REGION Network 12: Lowest Value of 2
   RUNG wire#powerrail
      Contact( #HMI.Alarms.oneTxFaulted )
      I_Contact( #HMI.Alarms.twoTxFaulted )
      { S7_Templates := "SrcType := Int" } EQ_Contact(in1 := #HMI.Control.failMode, in2 := 7)
      Move(in := #lowest, out1 => #activeValue)
   END_RUNG
   // the same network as SCL:
   IF #HMI.Alarms.oneTxFaulted AND NOT #HMI.Alarms.twoTxFaulted AND (#HMI.Control.failMode = 7) THEN
       #activeValue := #lowest;
   END_IF;
END_REGION

REGION Network 13: Average Value
   RUNG wire#powerrail
      Contact( #fault3 )
      { S7_Templates := "SrcType := Real"; S7_Expression := "(IN1+IN2)/IN3" } Calculate(in1 := #analog1, in2 := #analog2, in3 := 2.0, out => #average)
   END_RUNG
   RUNG wire#powerrail
      Contact( #fault2 )
      { S7_Templates := "SrcType := Real"; S7_Expression := "(IN1+IN2)/IN3" } Calculate(in1 := #analog1, in2 := #analog3, in3 := 2.0, out => #average)
   END_RUNG
   RUNG wire#powerrail
      Contact( #fault1 )
      { S7_Templates := "SrcType := Real"; S7_Expression := "(IN1+IN2)/IN3" } Calculate(in1 := #analog3, in2 := #analog2, in3 := 2.0, out => #average)
   END_RUNG
   RUNG wire#powerrail
      I_Contact( #fault1 )
      I_Contact( #fault2 )
      I_Contact( #fault3 )
      { S7_Templates := "SrcType := Real"; S7_Expression := "(IN1+IN2+IN3)/IN4" } Calculate(in1 := #analog1, in2 := #analog2, in3 := #analog3, in4 := 3.0, out => #average)
   END_RUNG
   // the same network as SCL:
   IF #fault3 THEN #average := (#analog1+#analog2)/2.0; END_IF;
   IF #fault2 THEN #average := (#analog1+#analog3)/2.0; END_IF;
   IF #fault1 THEN #average := (#analog3+#analog2)/2.0; END_IF;
   IF NOT #fault1 AND NOT #fault2 AND NOT #fault3 THEN #average := (#analog1+#analog2+#analog3)/3.0; END_IF;
END_REGION

REGION Network 14: Average of 3 values
   RUNG wire#powerrail
      { S7_Templates := "SrcType := Int" } EQ_Contact(in1 := #HMI.Control.mode, in2 := 4)
      wire#w1
      Move(in := #average, out1 => #activeValue)
   END_RUNG
   RUNG wire#powerrail
      Contact( #HMI.Alarms.oneTxFaulted )
      I_Contact( #HMI.Alarms.twoTxFaulted )
      { S7_Templates := "SrcType := Int" } EQ_Contact(in1 := #HMI.Control.failMode, in2 := 4)
   END_RUNG wire#w1
   // the same network as SCL:
   IF (#HMI.Control.mode = 4) OR (#HMI.Alarms.oneTxFaulted AND NOT #HMI.Alarms.twoTxFaulted AND (#HMI.Control.failMode = 4)) THEN
       #activeValue := #average;
   END_IF;
END_REGION

REGION Network 15: HH Voting Value 1
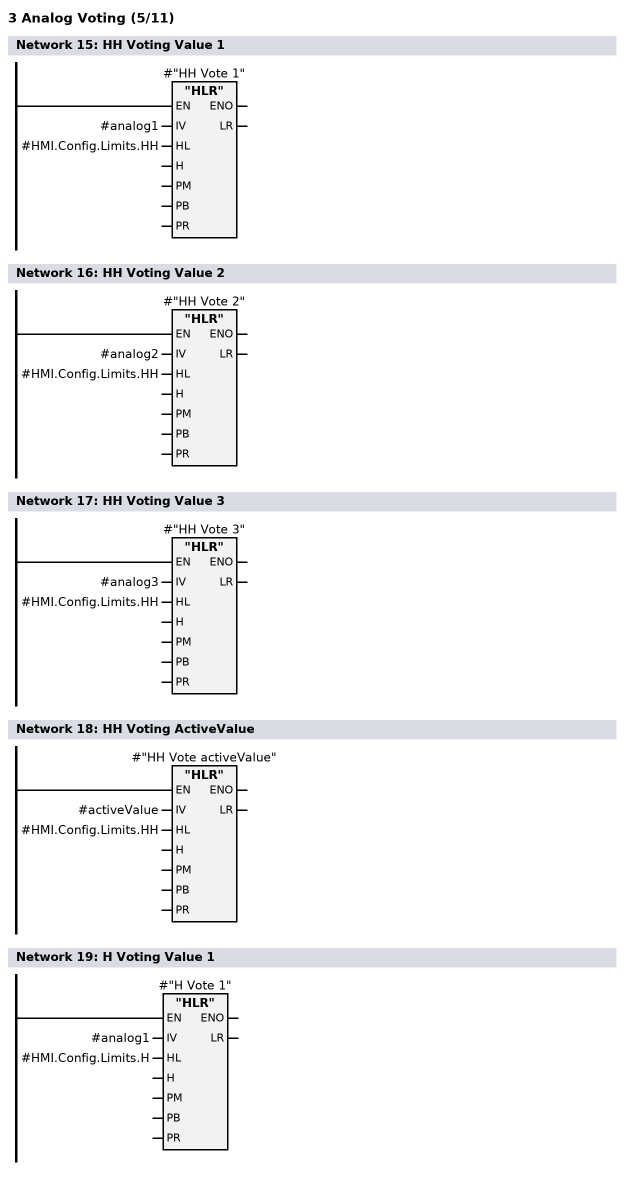
   RUNG wire#powerrail
      #"HH Vote 1"(IV := #analog1, HL := #HMI.Config.Limits.HH, H :=, PM :=, PB :=, PR :=, LR =>)
   END_RUNG
   // the same network as SCL:
   #"HH Vote 1"(IV := #analog1, HL := #HMI.Config.Limits.HH);   // "HLR"
END_REGION

REGION Network 16: HH Voting Value 2
   RUNG wire#powerrail
      #"HH Vote 2"(IV := #analog2, HL := #HMI.Config.Limits.HH, H :=, PM :=, PB :=, PR :=, LR =>)
   END_RUNG
   // the same network as SCL:
   #"HH Vote 2"(IV := #analog2, HL := #HMI.Config.Limits.HH);   // "HLR"
END_REGION

REGION Network 17: HH Voting Value 3
   RUNG wire#powerrail
      #"HH Vote 3"(IV := #analog3, HL := #HMI.Config.Limits.HH, H :=, PM :=, PB :=, PR :=, LR =>)
   END_RUNG
   // the same network as SCL:
   #"HH Vote 3"(IV := #analog3, HL := #HMI.Config.Limits.HH);   // "HLR"
END_REGION

REGION Network 18: HH Voting ActiveValue
   RUNG wire#powerrail
      #"HH Vote activeValue"(IV := #activeValue, HL := #HMI.Config.Limits.HH, H :=, PM :=, PB :=, PR :=, LR =>)
   END_RUNG
   // the same network as SCL:
   #"HH Vote activeValue"(IV := #activeValue, HL := #HMI.Config.Limits.HH);   // "HLR"
END_REGION

REGION Network 19: H Voting Value 1
   RUNG wire#powerrail
      #"H Vote 1"(IV := #analog1, HL := #HMI.Config.Limits.H, H :=, PM :=, PB :=, PR :=, LR =>)
   END_RUNG
   // the same network as SCL:
   #"H Vote 1"(IV := #analog1, HL := #HMI.Config.Limits.H);   // "HLR"
END_REGION

REGION Network 20: H Voting Value 2
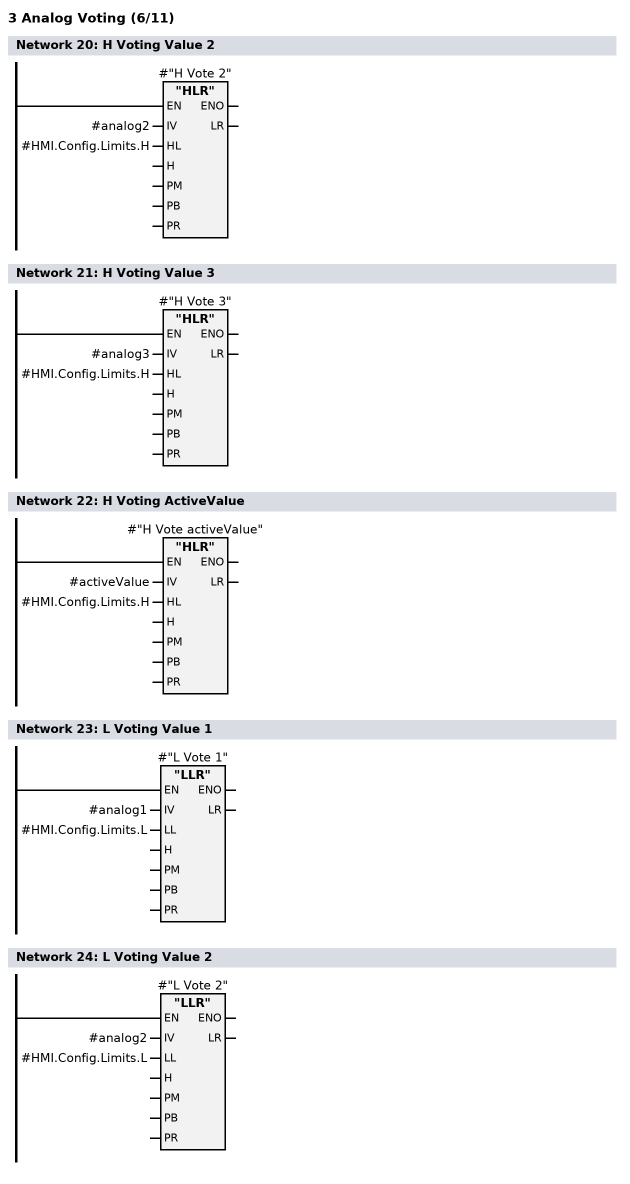
   RUNG wire#powerrail
      #"H Vote 2"(IV := #analog2, HL := #HMI.Config.Limits.H, H :=, PM :=, PB :=, PR :=, LR =>)
   END_RUNG
   // the same network as SCL:
   #"H Vote 2"(IV := #analog2, HL := #HMI.Config.Limits.H);   // "HLR"
END_REGION

REGION Network 21: H Voting Value 3
   RUNG wire#powerrail
      #"H Vote 3"(IV := #analog3, HL := #HMI.Config.Limits.H, H :=, PM :=, PB :=, PR :=, LR =>)
   END_RUNG
   // the same network as SCL:
   #"H Vote 3"(IV := #analog3, HL := #HMI.Config.Limits.H);   // "HLR"
END_REGION

REGION Network 22: H Voting ActiveValue
   RUNG wire#powerrail
      #"H Vote activeValue"(IV := #activeValue, HL := #HMI.Config.Limits.H, H :=, PM :=, PB :=, PR :=, LR =>)
   END_RUNG
   // the same network as SCL:
   #"H Vote activeValue"(IV := #activeValue, HL := #HMI.Config.Limits.H);   // "HLR"
END_REGION

REGION Network 23: L Voting Value 1
   RUNG wire#powerrail
      #"L Vote 1"(IV := #analog1, LL := #HMI.Config.Limits.L, H :=, PM :=, PB :=, PR :=, LR =>)
   END_RUNG
   // the same network as SCL:
   #"L Vote 1"(IV := #analog1, LL := #HMI.Config.Limits.L);   // "LLR"
END_REGION

REGION Network 24: L Voting Value 2
   RUNG wire#powerrail
      #"L Vote 2"(IV := #analog2, LL := #HMI.Config.Limits.L, H :=, PM :=, PB :=, PR :=, LR =>)
   END_RUNG
   // the same network as SCL:
   #"L Vote 2"(IV := #analog2, LL := #HMI.Config.Limits.L);   // "LLR"
END_REGION

REGION Network 25: L Voting Value 3
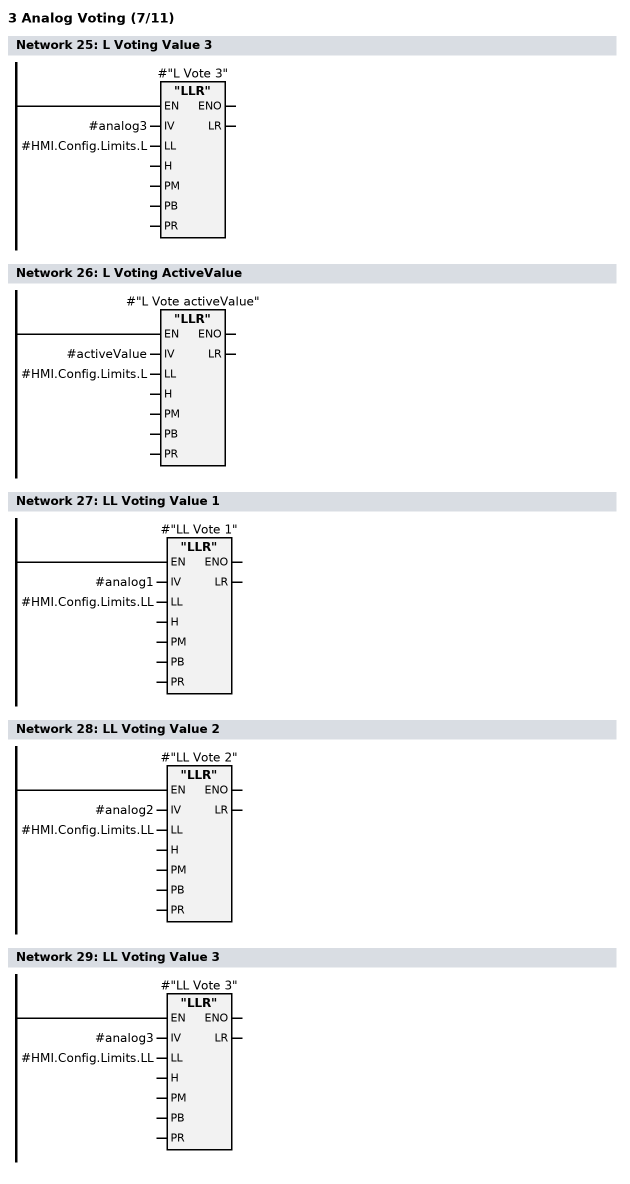
   RUNG wire#powerrail
      #"L Vote 3"(IV := #analog3, LL := #HMI.Config.Limits.L, H :=, PM :=, PB :=, PR :=, LR =>)
   END_RUNG
   // the same network as SCL:
   #"L Vote 3"(IV := #analog3, LL := #HMI.Config.Limits.L);   // "LLR"
END_REGION

REGION Network 26: L Voting ActiveValue
   RUNG wire#powerrail
      #"L Vote activeValue"(IV := #activeValue, LL := #HMI.Config.Limits.L, H :=, PM :=, PB :=, PR :=, LR =>)
   END_RUNG
   // the same network as SCL:
   #"L Vote activeValue"(IV := #activeValue, LL := #HMI.Config.Limits.L);   // "LLR"
END_REGION

REGION Network 27: LL Voting Value 1
   RUNG wire#powerrail
      #"LL Vote 1"(IV := #analog1, LL := #HMI.Config.Limits.LL, H :=, PM :=, PB :=, PR :=, LR =>)
   END_RUNG
   // the same network as SCL:
   #"LL Vote 1"(IV := #analog1, LL := #HMI.Config.Limits.LL);   // "LLR"
END_REGION

REGION Network 28: LL Voting Value 2
   RUNG wire#powerrail
      #"LL Vote 2"(IV := #analog2, LL := #HMI.Config.Limits.LL, H :=, PM :=, PB :=, PR :=, LR =>)
   END_RUNG
   // the same network as SCL:
   #"LL Vote 2"(IV := #analog2, LL := #HMI.Config.Limits.LL);   // "LLR"
END_REGION

REGION Network 29: LL Voting Value 3
   RUNG wire#powerrail
      #"LL Vote 3"(IV := #analog3, LL := #HMI.Config.Limits.LL, H :=, PM :=, PB :=, PR :=, LR =>)
   END_RUNG
   // the same network as SCL:
   #"LL Vote 3"(IV := #analog3, LL := #HMI.Config.Limits.LL);   // "LLR"
END_REGION

REGION Network 30: LL Voting ActiveValue
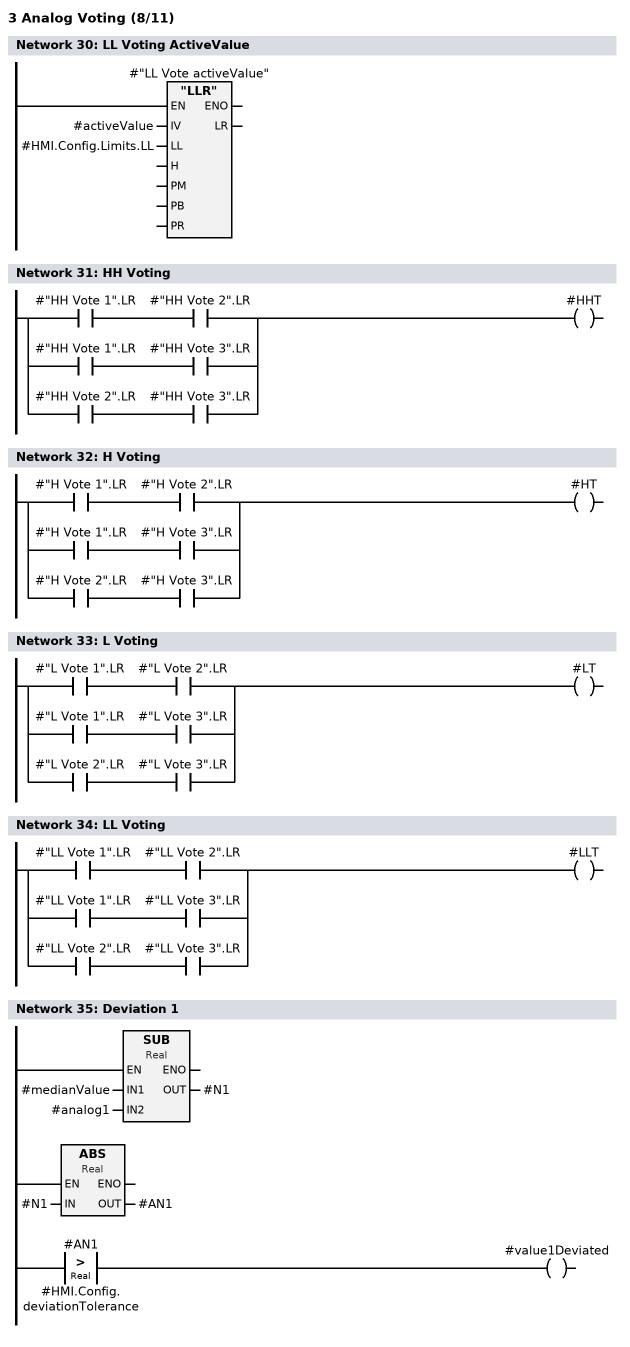
   RUNG wire#powerrail
      #"LL Vote activeValue"(IV := #activeValue, LL := #HMI.Config.Limits.LL, H :=, PM :=, PB :=, PR :=, LR =>)
   END_RUNG
   // the same network as SCL:
   #"LL Vote activeValue"(IV := #activeValue, LL := #HMI.Config.Limits.LL);   // "LLR"
END_REGION

REGION Network 31: HH Voting
   RUNG wire#powerrail
      Contact( #"HH Vote 1".LR )
      Contact( #"HH Vote 2".LR )
      wire#w1
      Coil( #HHT )
   END_RUNG
   RUNG wire#powerrail
      Contact( #"HH Vote 1".LR )
      Contact( #"HH Vote 3".LR )
   END_RUNG wire#w1
   RUNG wire#powerrail
      Contact( #"HH Vote 2".LR )
      Contact( #"HH Vote 3".LR )
   END_RUNG wire#w1
   // the same network as SCL:
   #HHT := (#"HH Vote 1".LR AND #"HH Vote 2".LR) OR (#"HH Vote 1".LR AND #"HH Vote 3".LR) OR (#"HH Vote 2".LR AND #"HH Vote 3".LR);
END_REGION

REGION Network 32: H Voting
   RUNG wire#powerrail
      Contact( #"H Vote 1".LR )
      Contact( #"H Vote 2".LR )
      wire#w1
      Coil( #HT )
   END_RUNG
   RUNG wire#powerrail
      Contact( #"H Vote 1".LR )
      Contact( #"H Vote 3".LR )
   END_RUNG wire#w1
   RUNG wire#powerrail
      Contact( #"H Vote 2".LR )
      Contact( #"H Vote 3".LR )
   END_RUNG wire#w1
   // the same network as SCL:
   #HT := (#"H Vote 1".LR AND #"H Vote 2".LR) OR (#"H Vote 1".LR AND #"H Vote 3".LR) OR (#"H Vote 2".LR AND #"H Vote 3".LR);
END_REGION

REGION Network 33: L Voting
   RUNG wire#powerrail
      Contact( #"L Vote 1".LR )
      Contact( #"L Vote 2".LR )
      wire#w1
      Coil( #LT )
   END_RUNG
   RUNG wire#powerrail
      Contact( #"L Vote 1".LR )
      Contact( #"L Vote 3".LR )
   END_RUNG wire#w1
   RUNG wire#powerrail
      Contact( #"L Vote 2".LR )
      Contact( #"L Vote 3".LR )
   END_RUNG wire#w1
   // the same network as SCL:
   #LT := (#"L Vote 1".LR AND #"L Vote 2".LR) OR (#"L Vote 1".LR AND #"L Vote 3".LR) OR (#"L Vote 2".LR AND #"L Vote 3".LR);
END_REGION

REGION Network 34: LL Voting
   RUNG wire#powerrail
      Contact( #"LL Vote 1".LR )
      Contact( #"LL Vote 2".LR )
      wire#w1
      Coil( #LLT )
   END_RUNG
   RUNG wire#powerrail
      Contact( #"LL Vote 1".LR )
      Contact( #"LL Vote 3".LR )
   END_RUNG wire#w1
   RUNG wire#powerrail
      Contact( #"LL Vote 2".LR )
      Contact( #"LL Vote 3".LR )
   END_RUNG wire#w1
   // the same network as SCL:
   #LLT := (#"LL Vote 1".LR AND #"LL Vote 2".LR) OR (#"LL Vote 1".LR AND #"LL Vote 3".LR) OR (#"LL Vote 2".LR AND #"LL Vote 3".LR);
END_REGION

REGION Network 35: Deviation 1
   RUNG wire#powerrail
      { S7_Templates := "SrcType := Real"; S7_GenerateENO := "TRUE" } Sub(in1 := #medianValue, in2 := #analog1, out => #N1)
   END_RUNG
   RUNG wire#powerrail
      { S7_Templates := "SrcType := Real"; S7_GenerateENO := "TRUE" } Abs(in := #N1, out => #AN1)
   END_RUNG
   RUNG wire#powerrail
      { S7_Templates := "SrcType := Real" } GT_Contact(in1 := #AN1, in2 := #HMI.Config.deviationTolerance)
      Coil( #value1Deviated )
   END_RUNG
   // the same network as SCL:
   #N1 := #medianValue - #analog1;
   #AN1 := ABS(#N1);
   #value1Deviated := #AN1 > #HMI.Config.deviationTolerance;
END_REGION

REGION Network 36: Deviation 2
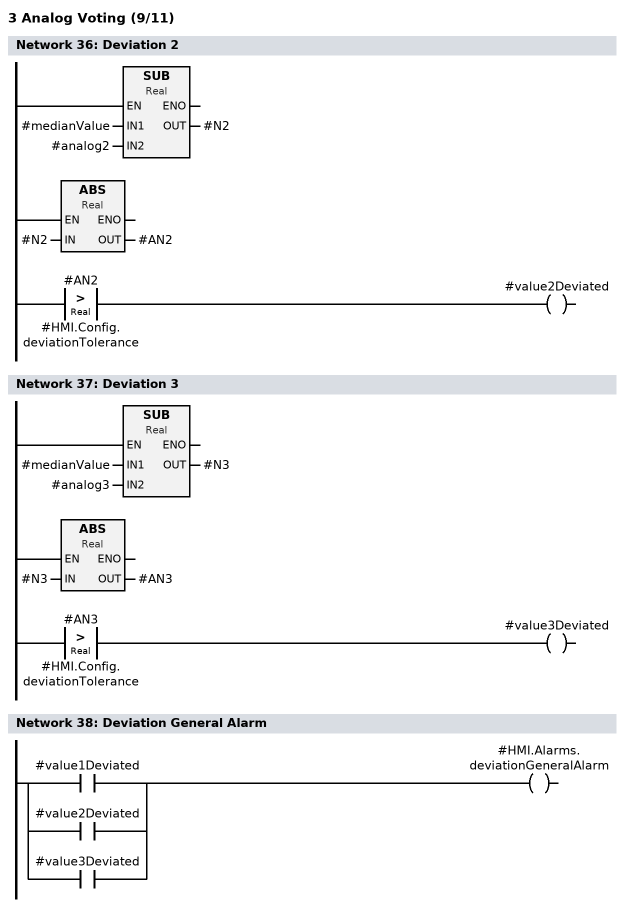
   RUNG wire#powerrail
      { S7_Templates := "SrcType := Real"; S7_GenerateENO := "TRUE" } Sub(in1 := #medianValue, in2 := #analog2, out => #N2)
   END_RUNG
   RUNG wire#powerrail
      { S7_Templates := "SrcType := Real"; S7_GenerateENO := "TRUE" } Abs(in := #N2, out => #AN2)
   END_RUNG
   RUNG wire#powerrail
      { S7_Templates := "SrcType := Real" } GT_Contact(in1 := #AN2, in2 := #HMI.Config.deviationTolerance)
      Coil( #value2Deviated )
   END_RUNG
   // the same network as SCL:
   #N2 := #medianValue - #analog2;
   #AN2 := ABS(#N2);
   #value2Deviated := #AN2 > #HMI.Config.deviationTolerance;
END_REGION

REGION Network 37: Deviation 3
   RUNG wire#powerrail
      { S7_Templates := "SrcType := Real"; S7_GenerateENO := "TRUE" } Sub(in1 := #medianValue, in2 := #analog3, out => #N3)
   END_RUNG
   RUNG wire#powerrail
      { S7_Templates := "SrcType := Real"; S7_GenerateENO := "TRUE" } Abs(in := #N3, out => #AN3)
   END_RUNG
   RUNG wire#powerrail
      { S7_Templates := "SrcType := Real" } GT_Contact(in1 := #AN3, in2 := #HMI.Config.deviationTolerance)
      Coil( #value3Deviated )
   END_RUNG
   // the same network as SCL:
   #N3 := #medianValue - #analog3;
   #AN3 := ABS(#N3);
   #value3Deviated := #AN3 > #HMI.Config.deviationTolerance;
END_REGION

REGION Network 38: Deviation General Alarm
   RUNG wire#powerrail
      Contact( #value1Deviated )
      wire#w1
      Coil( #HMI.Alarms.deviationGeneralAlarm )
   END_RUNG
   RUNG wire#powerrail
      Contact( #value2Deviated )
   END_RUNG wire#w1
   RUNG wire#powerrail
      Contact( #value3Deviated )
   END_RUNG wire#w1
   // the same network as SCL:
   #HMI.Alarms.deviationGeneralAlarm := #value1Deviated OR #value2Deviated OR #value3Deviated;
END_REGION

REGION Network 39: Master Trip
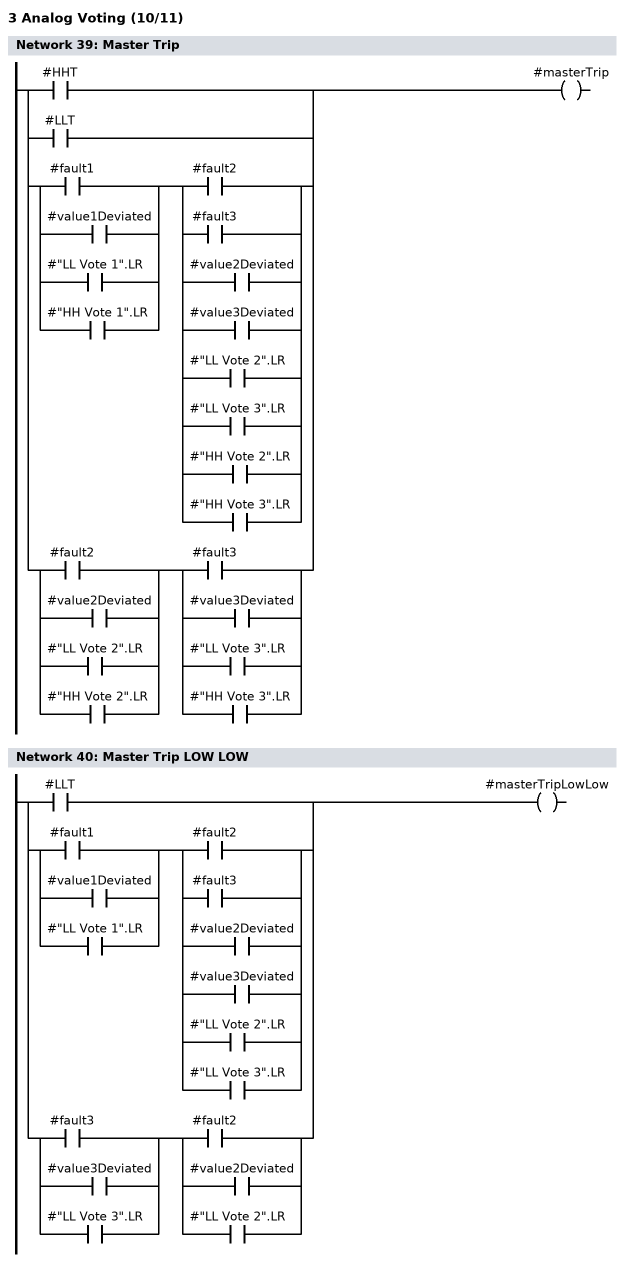
   RUNG wire#powerrail
      Contact( #HHT )
      wire#w1
      Coil( #masterTrip )
   END_RUNG
   RUNG wire#powerrail
      Contact( #LLT )
   END_RUNG wire#w1
   RUNG wire#powerrail
      Contact( #fault1 )
      wire#w2
      Contact( #fault2 )
   END_RUNG wire#w1
   RUNG wire#powerrail
      Contact( #value1Deviated )
   END_RUNG wire#w2
   RUNG wire#powerrail
      Contact( #"LL Vote 1".LR )
   END_RUNG wire#w2
   RUNG wire#powerrail
      Contact( #"HH Vote 1".LR )
   END_RUNG wire#w2
   RUNG wire#w2
      Contact( #fault3 )
   END_RUNG wire#w1
   RUNG wire#w2
      Contact( #value2Deviated )
   END_RUNG wire#w1
   RUNG wire#w2
      Contact( #value3Deviated )
   END_RUNG wire#w1
   RUNG wire#w2
      Contact( #"LL Vote 2".LR )
   END_RUNG wire#w1
   RUNG wire#w2
      Contact( #"LL Vote 3".LR )
   END_RUNG wire#w1
   RUNG wire#w2
      Contact( #"HH Vote 2".LR )
   END_RUNG wire#w1
   RUNG wire#w2
      Contact( #"HH Vote 3".LR )
   END_RUNG wire#w1
   RUNG wire#powerrail
      Contact( #fault2 )
      wire#w3
      Contact( #fault3 )
   END_RUNG wire#w1
   RUNG wire#powerrail
      Contact( #value2Deviated )
   END_RUNG wire#w3
   RUNG wire#powerrail
      Contact( #"LL Vote 2".LR )
   END_RUNG wire#w3
   RUNG wire#powerrail
      Contact( #"HH Vote 2".LR )
   END_RUNG wire#w3
   RUNG wire#w3
      Contact( #value3Deviated )
   END_RUNG wire#w1
   RUNG wire#w3
      Contact( #"LL Vote 3".LR )
   END_RUNG wire#w1
   RUNG wire#w3
      Contact( #"HH Vote 3".LR )
   END_RUNG wire#w1
   // the same network as SCL:
   #masterTrip := #HHT OR #LLT OR ((#fault1 OR #value1Deviated OR #"LL Vote 1".LR OR #"HH Vote 1".LR) AND (#fault2 OR #fault3 OR #value2Deviated OR #value3Deviated OR #"LL Vote 2".LR OR #"LL Vote 3".LR OR #"HH Vote 2".LR OR #"HH Vote 3".LR)) OR ((#fault2 OR #value2Deviated OR #"LL Vote 2".LR OR #"HH Vote 2".LR) AND (#fault3 OR #value3Deviated OR #"LL Vote 3".LR OR #"HH Vote 3".LR));
END_REGION

REGION Network 40: Master Trip LOW LOW
   RUNG wire#powerrail
      Contact( #LLT )
      wire#w1
      Coil( #masterTripLowLow )
   END_RUNG
   RUNG wire#powerrail
      Contact( #fault1 )
      wire#w2
      Contact( #fault2 )
   END_RUNG wire#w1
   RUNG wire#powerrail
      Contact( #value1Deviated )
   END_RUNG wire#w2
   RUNG wire#powerrail
      Contact( #"LL Vote 1".LR )
   END_RUNG wire#w2
   RUNG wire#w2
      Contact( #fault3 )
   END_RUNG wire#w1
   RUNG wire#w2
      Contact( #value2Deviated )
   END_RUNG wire#w1
   RUNG wire#w2
      Contact( #value3Deviated )
   END_RUNG wire#w1
   RUNG wire#w2
      Contact( #"LL Vote 2".LR )
   END_RUNG wire#w1
   RUNG wire#w2
      Contact( #"LL Vote 3".LR )
   END_RUNG wire#w1
   RUNG wire#powerrail
      Contact( #fault3 )
      wire#w3
      Contact( #fault2 )
   END_RUNG wire#w1
   RUNG wire#powerrail
      Contact( #value3Deviated )
   END_RUNG wire#w3
   RUNG wire#powerrail
      Contact( #"LL Vote 3".LR )
   END_RUNG wire#w3
   RUNG wire#w3
      Contact( #value2Deviated )
   END_RUNG wire#w1
   RUNG wire#w3
      Contact( #"LL Vote 2".LR )
   END_RUNG wire#w1
   // the same network as SCL:
   #masterTripLowLow := #LLT OR ((#fault1 OR #value1Deviated OR #"LL Vote 1".LR) AND (#fault2 OR #fault3 OR #value2Deviated OR #value3Deviated OR #"LL Vote 2".LR OR #"LL Vote 3".LR)) OR ((#fault3 OR #value3Deviated OR #"LL Vote 3".LR) AND (#fault2 OR #value2Deviated OR #"LL Vote 2".LR));
END_REGION

REGION Network 41: Master Trip HIGH HIGH
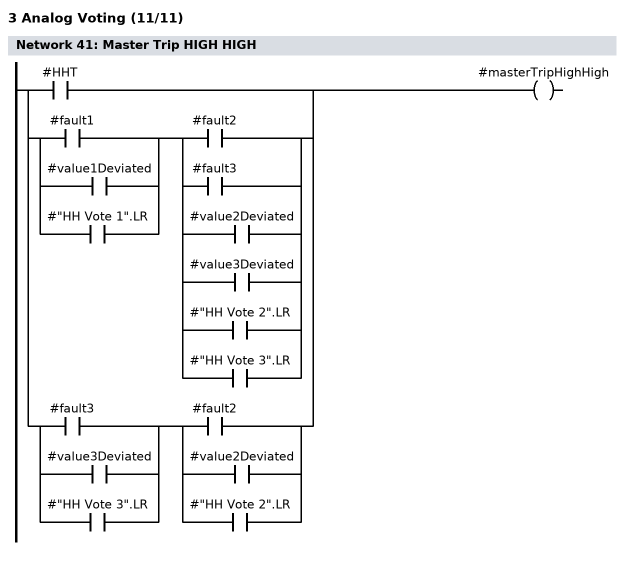
   RUNG wire#powerrail
      Contact( #HHT )
      wire#w1
      Coil( #masterTripHighHigh )
   END_RUNG
   RUNG wire#powerrail
      Contact( #fault1 )
      wire#w2
      Contact( #fault2 )
   END_RUNG wire#w1
   RUNG wire#powerrail
      Contact( #value1Deviated )
   END_RUNG wire#w2
   RUNG wire#powerrail
      Contact( #"HH Vote 1".LR )
   END_RUNG wire#w2
   RUNG wire#w2
      Contact( #fault3 )
   END_RUNG wire#w1
   RUNG wire#w2
      Contact( #value2Deviated )
   END_RUNG wire#w1
   RUNG wire#w2
      Contact( #value3Deviated )
   END_RUNG wire#w1
   RUNG wire#w2
      Contact( #"HH Vote 2".LR )
   END_RUNG wire#w1
   RUNG wire#w2
      Contact( #"HH Vote 3".LR )
   END_RUNG wire#w1
   RUNG wire#powerrail
      Contact( #fault3 )
      wire#w3
      Contact( #fault2 )
   END_RUNG wire#w1
   RUNG wire#powerrail
      Contact( #value3Deviated )
   END_RUNG wire#w3
   RUNG wire#powerrail
      Contact( #"HH Vote 3".LR )
   END_RUNG wire#w3
   RUNG wire#w3
      Contact( #value2Deviated )
   END_RUNG wire#w1
   RUNG wire#w3
      Contact( #"HH Vote 2".LR )
   END_RUNG wire#w1
   // the same network as SCL:
   #masterTripHighHigh := #HHT OR ((#fault1 OR #value1Deviated OR #"HH Vote 1".LR) AND (#fault2 OR #fault3 OR #value2Deviated OR #value3Deviated OR #"HH Vote 2".LR OR #"HH Vote 3".LR)) OR ((#fault3 OR #value3Deviated OR #"HH Vote 3".LR) AND (#fault2 OR #value2Deviated OR #"HH Vote 2".LR));
END_REGION
END_FUNCTION_BLOCK

FUNCTION_BLOCK "TX-AI"   // FB804, LAD
TITLE = SSAC Analog Trasmitter Function Block
{ S7_Optimized_Access := 'TRUE' }
VERSION : 1.0
// Default mode 0 starts at  network 6
   VAR_INPUT
      Mode : Int;   // TX Mode - 0 = 4-20 mA / 1 = Int Math (RTD/TC) / 2 = Real Input Conversion / 3 = SQRT / 5 = Simulated Transmitter Value / 6 = Vortex Flow Transmitters
      RAIVI : Int;   // Raw Analog Input Value INT
      RAIVR : Real;   // Raw Analog Input Value REAL
      EnableHighAlarms : Bool := True;
      EnableLowAlarms : Bool := True;
      "TI Fail" : Bool;
   END_VAR
   VAR_OUTPUT
      SAI : Real;   // Compensated Scaled Analog Value
   END_VAR
   VAR
      HMI : Struct   // Alarms
         Status : Struct
            USAV : Real;   // Uncompensated Scaled Analog Value
            TCV : Real;   // Temperature Compensation Value
            PCV : Real;   // Pressure Compensation Value
            NV : Real;   // Normalized Value
         END_STRUCT;
         Alarm : Struct
            Alarms : Word;
         END_STRUCT;
         Diag : Struct   // Diagnostics
            SV : Real;   // Simulation Value
         END_STRUCT;
      END_STRUCT;
   END_VAR
   VAR RETAIN
      Retain : Struct
         HMI : Struct
            Config : Struct   // Settings
               RIMXV : Real := 27648.0;   // Raw Input Maximum Value (Used for Sqrt)
               RIMNV : Real;   // Raw Input Minimum Value (Used for Sqrt)
               ESMXV : Real := 100.0;   // Engineering/Scaled Maximum Value
               ESMNV : Real;   // Engineering/Scaled Minimum Value
               COV : Bool;   // Clamp Output Value
               OV : Real;   // Offset Value
               SAM : Bool;   // Substitution Activation Mode
               SAV : Real := -999999.0;   // Substitution Value during a limit input value trip
               CE : Struct   // Compensation Equation
                  TC : Real := 460.0;   // Temperature Constant
                  PC : Real := 14.7;   // Pressure Constant
                  TR : Real := 1.0;   // Temperature Reference
                  TA : Real := 1.0;   // Temperature Actual
                  PR : Real := 1.0;   // Pressure Reference
                  PA : Real := 1.0;   // Pressure Actual
               END_STRUCT;
               SP : Struct   // Setpoints
                  Limits : Struct
                     HHH : Real := 95.0;   // HHH Limit Setpoint
                     HH : Real := 90.0;   // HH Limit Setpoint
                     H : Real := 80.0;   // HH Limit Setpoint
                     L : Real := 20.0;   // L Limit Setpoint
                     LL : Real := 10.0;   // LL Limit Setpoint
                     LLL : Real := 5.0;   // LLL Limit Setpoint
                     "OR" : Real := 5.0;   // Over range value
                     UR : Real := 5.0;   // Under range value
                  END_STRUCT;
                  HYS : Struct   // Hysteresis
                     Global : Real;   // Hysteresis global value, only valid when greater than or equal to 0
                     HHH : Real := 1.0;   // Hysteresis Setpoint - High High High
                     HH : Real := 1.0;   // Hysteresis Setpoint - High High
                     H : Real := 1.0;   // Hysteresis Setpoint - High
                     L : Real := 1.0;   // Hysteresis Setpoint - Low
                     LL : Real := 1.0;   // Hysteresis Setpoint - Low Low
                     LLL : Real := 1.0;   // Hysteresis Setpoint - Low Low Low
                     "OR" : Real := 1.0;   // Hysteresis Setpoint - Over Range
                     UR : Real := 1.0;   // Hysteresis Setpoint - Under Range
                  END_STRUCT;
                  SUB_ON : Bool;   // Substitution Activation
               END_STRUCT;
               PT : Struct   // Setpoints
                  HLD : Struct   // Hold
                     Global : Time;   // Hold PT global value, only valid when not equal to 0
                     AHHH : Time := t#5s;   // Alarm Debounce
                     AHH : Time := t#5s;   // Alarm Debounce
                     AH : Time := t#5s;   // Alarm Debounce
                     AL : Time := t#5s;   // Alarm Debounce
                     ALL : Time := t#5s;   // Alarm Debounce
                     ALLL : Time := t#5s;   // Alarm Debounce
                     "OR" : Time := t#5s;   // Over range hold
                     UR : Time := t#5s;   // Under range hold
                  END_STRUCT;
                  DBNC : Struct   // Debounce
                     Global : Time;   // Debounce PT global value, only valid when not equal to 0
                     AHHH : Time := t#5s;   // Alarm Debounce
                     AHH : Time := t#5s;   // Alarm Debounce
                     AH : Time := t#5s;   // Alarm Debounce
                     AL : Time := t#5s;   // Alarm Debounce
                     ALL : Time := t#5s;   // Alarm Debounce
                     ALLL : Time := t#5s;   // Alarm Debounce
                     "OR" : Time := t#5s;   // Over range debounce
                     UR : Time := t#5s;   // Under range debounce
                  END_STRUCT;
               END_STRUCT;
               Alarms : Word := 16#01FF;
            END_STRUCT;
         END_STRUCT;
      END_STRUCT;
   END_VAR
   VAR
      Admin : Struct   // Admin configurations
         SCL : Struct   // Scale Values
            RDP : Real := 10.0;   // RTD Decimal Places
            RRIMD : Real := 1.0;   // Raw Real input Math divider
            "OR" : Real;   // Over Range Value
            UR : Real;   // Under Range Value
            SAIV : Real;   // Scaled Analog Input Value
         END_STRUCT;
         HYS : Struct   // Hysteresis - Computed Values
            "OR" : Real;   // Hysteresis Value - Over Range
            UR : Real;   // Hysteresis Value - Under Range
         END_STRUCT;
      END_STRUCT;
      Alarms : Struct
         HighHighHigh : Bool;
         HighHigh : Bool;
         High : Bool;
         Low : Bool;
         LowLow : Bool;
         LowLowLow : Bool;
         TransmitterFault : Bool;
         UnderRange : Bool;
         OverRange : Bool;
      END_STRUCT;
      Timers : Struct
         OR_DB : TON_TIME;   // Over Range Debounce
         UR_DB : TON_TIME;   // Under Range DB
         OR_HLD : TOF_TIME;   // Over Range Hold
         UR_HLD : TOF_TIME;   // Under Range Hold
         DBNC : Struct
            HHH : TON_TIME;
            HH : TON_TIME;
            H : TON_TIME;
            L : TON_TIME;
            LL : TON_TIME;
            LLL : TON_TIME;
         END_STRUCT;
         HOLD : Struct
            HHH : TOF_TIME;
            HH : TOF_TIME;
            H : TOF_TIME;
            L : TOF_TIME;
            LL : TOF_TIME;
            LLL : TOF_TIME;
         END_STRUCT;
      END_STRUCT;
      molActual : Real := 1.0;
      molDesign : Real := 1.0;
   END_VAR
   VAR_TEMP
      SRV : Real;
      RAIDI : DInt;   // Raw Analog Input DINT
      RAIR : Real;   // Raw Analog Input REAL
      RAIAV : Real;   // Raw Analog Input Absolute Value
      RAIVS : Real;   // Raw Analog Input Value Scaler
      TCRE : Real;   // Temperature Compensation Reference Equation
      TCAE : Real;   // Temperature Compensation Actual Equation
      PCRE : Real;   // Pressure Compensation Reference Equation
      PCAE : Real;   // Pressure Compensation Actual Equation
      TPCV : Real;   // Temperature Pressure Compensation Value
      MWCV : Real;   // Mol Weight Compensation Value
      TPMCV : Real;   // Temperature Pressure Mol Compensation Value
      sqrtSaiv : Real;   // SCALED ANALOG INT VALUE TO BE SQRT'D
      rawValue : Int;
      dummy : Bool;
      sqrt01 : Real;
      RAIVR_1 : DInt;
      RAIVR_1_1 : Real;
      ValuePerPoint : Real;
      ValueAddRaw : Real;
      "DBNC.SP" : Struct
         HHH : Real;
         HH : Real;
         H : Real;
         L : Real;
         LL : Real;
         LLL : Real;
      END_STRUCT;
   END_VAR
   VAR_TEMP   // added for the SCL form of the ladder/FBD networks
      _w1 : Bool;
      _w2 : Bool;
   END_VAR
BEGIN

REGION Network 1: Transmitter Mode 1 = Int Math or RTD
   // MD1 Jump to network 9
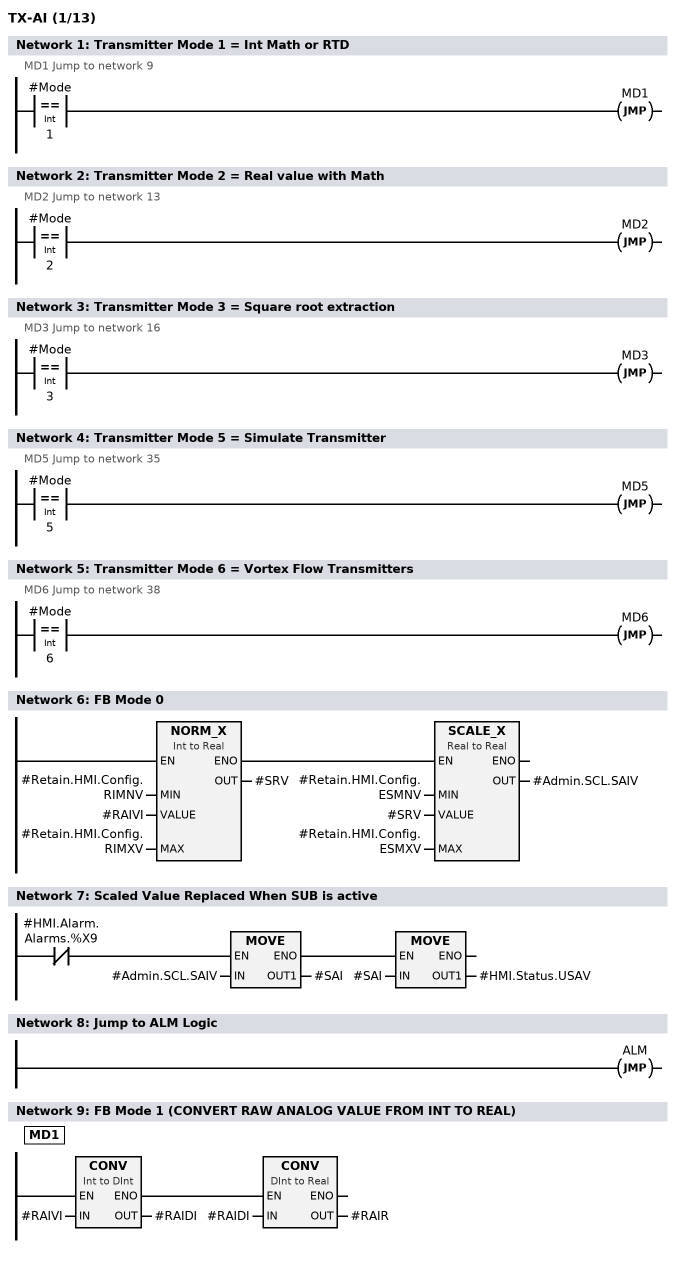
   RUNG wire#powerrail
      { S7_Templates := "SrcType := Int" } EQ_Contact(in1 := #Mode, in2 := 1)
      JumpCoil( MD1 )
   END_RUNG
   // the same network as SCL:
   IF #Mode = 1 THEN GOTO MD1; END_IF;
END_REGION

REGION Network 2: Transmitter Mode 2 = Real value with Math
   // MD2 Jump to network 13
   RUNG wire#powerrail
      { S7_Templates := "SrcType := Int" } EQ_Contact(in1 := #Mode, in2 := 2)
      JumpCoil( MD2 )
   END_RUNG
   // the same network as SCL:
   IF #Mode = 2 THEN GOTO MD2; END_IF;
END_REGION

REGION Network 3: Transmitter Mode 3 = Square root extraction
   // MD3 Jump to network 16
   RUNG wire#powerrail
      { S7_Templates := "SrcType := Int" } EQ_Contact(in1 := #Mode, in2 := 3)
      JumpCoil( MD3 )
   END_RUNG
   // the same network as SCL:
   IF #Mode = 3 THEN GOTO MD3; END_IF;
END_REGION

REGION Network 4: Transmitter Mode 5 = Simulate Transmitter
   // MD5 Jump to network 35
   RUNG wire#powerrail
      { S7_Templates := "SrcType := Int" } EQ_Contact(in1 := #Mode, in2 := 5)
      JumpCoil( MD5 )
   END_RUNG
   // the same network as SCL:
   IF #Mode = 5 THEN GOTO MD5; END_IF;
END_REGION

REGION Network 5: Transmitter Mode 6 = Vortex Flow Transmitters
   // MD6 Jump to network 38
   RUNG wire#powerrail
      { S7_Templates := "SrcType := Int" } EQ_Contact(in1 := #Mode, in2 := 6)
      JumpCoil( MD6 )
   END_RUNG
   // the same network as SCL:
   IF #Mode = 6 THEN GOTO MD6; END_IF;
END_REGION

REGION Network 6: FB Mode 0
   RUNG wire#powerrail
      { S7_Templates := "[SrcType := Int, DestType := Real]" } Normalize(min := #Retain.HMI.Config.RIMNV, value := #RAIVI, max := #Retain.HMI.Config.RIMXV, out => #SRV)
      { S7_Templates := "[SrcType := Real, DestType := Real]" } Scale(min := #Retain.HMI.Config.ESMNV, value := #SRV, max := #Retain.HMI.Config.ESMXV, out => #Admin.SCL.SAIV)
   END_RUNG
   // the same network as SCL:
   #SRV := NORM_X(MIN := #Retain.HMI.Config.RIMNV, VALUE := #RAIVI, MAX := #Retain.HMI.Config.RIMXV);
   #Admin.SCL.SAIV := SCALE_X(MIN := #Retain.HMI.Config.ESMNV, VALUE := #SRV, MAX := #Retain.HMI.Config.ESMXV);
END_REGION

REGION Network 7: Scaled Value Replaced When SUB is active
   RUNG wire#powerrail
      I_Contact( #HMI.Alarm.Alarms.%X9 )
      { S7_GenerateENO := "TRUE" } Move(in := #Admin.SCL.SAIV, out1 => #SAI)
      { S7_GenerateENO := "TRUE" } Move(in := #SAI, out1 => #HMI.Status.USAV)
   END_RUNG
   // the same network as SCL:
   // ENO of a box is taken as its EN; it also drops when the box reports an error
   IF NOT #HMI.Alarm.Alarms.%X9 THEN
       #SAI := #Admin.SCL.SAIV;
       #HMI.Status.USAV := #SAI;
   END_IF;
END_REGION

REGION Network 8: Jump to ALM Logic
   RUNG wire#powerrail
      JumpCoil( ALM )
   END_RUNG
   // the same network as SCL:
   GOTO ALM;
END_REGION

REGION Network 9: FB Mode 1 (CONVERT RAW ANALOG VALUE FROM INT TO REAL)
   Label( MD1 )
   RUNG wire#powerrail
      { S7_Templates := "[SrcType := Int, DestType := DInt]"; S7_GenerateENO := "TRUE" } Convert(in := #RAIVI, out => #RAIDI)
      { S7_Templates := "[SrcType := DInt, DestType := Real]"; S7_GenerateENO := "TRUE" } Convert(in := #RAIDI, out => #RAIR)
   END_RUNG
   // the same network as SCL:
   // ENO of a box is taken as its EN; it also drops when the box reports an error
   MD1:
   #RAIDI := INT_TO_DINT(#RAIVI);
   #RAIR := DINT_TO_REAL(#RAIDI);
END_REGION

REGION Network 10: Raw RTD/TC value scaled based on divider
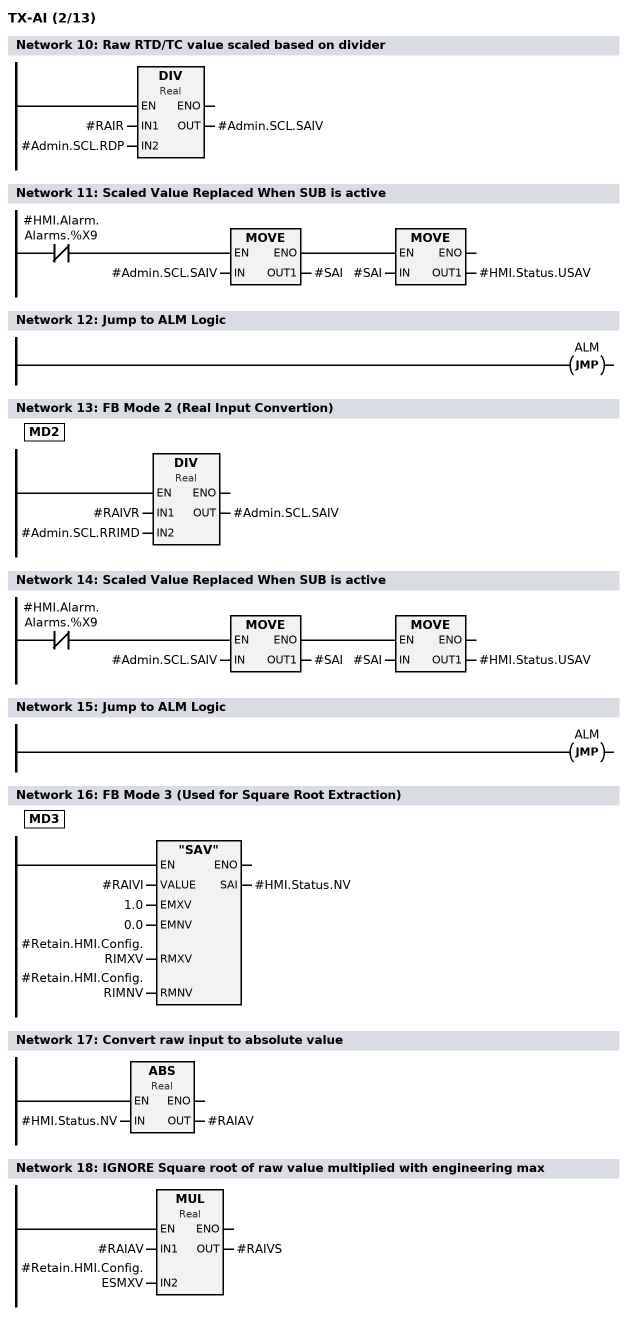
   RUNG wire#powerrail
      { S7_Templates := "SrcType := Real"; S7_GenerateENO := "TRUE" } Div(in1 := #RAIR, in2 := #Admin.SCL.RDP, out => #Admin.SCL.SAIV)
   END_RUNG
   // the same network as SCL:
   #Admin.SCL.SAIV := #RAIR / #Admin.SCL.RDP;
END_REGION

REGION Network 11: Scaled Value Replaced When SUB is active
   RUNG wire#powerrail
      I_Contact( #HMI.Alarm.Alarms.%X9 )
      { S7_GenerateENO := "TRUE" } Move(in := #Admin.SCL.SAIV, out1 => #SAI)
      Move(in := #SAI, out1 => #HMI.Status.USAV)
   END_RUNG
   // the same network as SCL:
   // ENO of a box is taken as its EN; it also drops when the box reports an error
   IF NOT #HMI.Alarm.Alarms.%X9 THEN
       #SAI := #Admin.SCL.SAIV;
       #HMI.Status.USAV := #SAI;
   END_IF;
END_REGION

REGION Network 12: Jump to ALM Logic
   RUNG wire#powerrail
      JumpCoil( ALM )
   END_RUNG
   // the same network as SCL:
   GOTO ALM;
END_REGION

REGION Network 13: FB Mode 2 (Real Input Convertion)
   Label( MD2 )
   RUNG wire#powerrail
      { S7_Templates := "SrcType := Real"; S7_GenerateENO := "TRUE" } Div(in1 := #RAIVR, in2 := #Admin.SCL.RRIMD, out => #Admin.SCL.SAIV)
   END_RUNG
   // the same network as SCL:
   MD2:
   #Admin.SCL.SAIV := #RAIVR / #Admin.SCL.RRIMD;
END_REGION

REGION Network 14: Scaled Value Replaced When SUB is active
   RUNG wire#powerrail
      I_Contact( #HMI.Alarm.Alarms.%X9 )
      { S7_GenerateENO := "TRUE" } Move(in := #Admin.SCL.SAIV, out1 => #SAI)
      Move(in := #SAI, out1 => #HMI.Status.USAV)
   END_RUNG
   // the same network as SCL:
   // ENO of a box is taken as its EN; it also drops when the box reports an error
   IF NOT #HMI.Alarm.Alarms.%X9 THEN
       #SAI := #Admin.SCL.SAIV;
       #HMI.Status.USAV := #SAI;
   END_IF;
END_REGION

REGION Network 15: Jump to ALM Logic
   RUNG wire#powerrail
      JumpCoil( ALM )
   END_RUNG
   // the same network as SCL:
   GOTO ALM;
END_REGION

REGION Network 16: FB Mode 3 (Used for Square Root Extraction)
   Label( MD3 )
   RUNG wire#powerrail
      "SAV"(VALUE := #RAIVI, EMXV := 1.0, EMNV := 0.0, RMXV := #Retain.HMI.Config.RIMXV, RMNV := #Retain.HMI.Config.RIMNV, SAI => #HMI.Status.NV)
   END_RUNG
   // the same network as SCL:
   MD3:
   "SAV"(VALUE := #RAIVI,
         EMXV := 1.0,
         EMNV := 0.0,
         RMXV := #Retain.HMI.Config.RIMXV,
         RMNV := #Retain.HMI.Config.RIMNV,
         SAI => #HMI.Status.NV);
END_REGION

REGION Network 17: Convert raw input to absolute value
   RUNG wire#powerrail
      { S7_Templates := "SrcType := Real"; S7_GenerateENO := "TRUE" } Abs(in := #HMI.Status.NV, out => #RAIAV)
   END_RUNG
   // the same network as SCL:
   #RAIAV := ABS(#HMI.Status.NV);
END_REGION

REGION Network 18: IGNORE Square root of raw value multiplied with engineering max
   RUNG wire#powerrail
      { S7_Templates := "SrcType := Real"; S7_GenerateENO := "TRUE" } Mul(in1 := #RAIAV, in2 := #Retain.HMI.Config.ESMXV, out => #RAIVS)
   END_RUNG
   // the same network as SCL:
   #RAIVS := #RAIAV * #Retain.HMI.Config.ESMXV;
END_REGION

REGION Network 19: Normalized Value greater than or equal to 0 move RAIVS into HMI.Status.USAV